
       REGION "COPY TO LOCAL"
           #selStnCount := #settings.current.stations.selCount;
       END_REGION

       REGION "ON CHANGE IN BUTTON OR STATION SELECTON"
           IF #settings.current.kp8.btnSelState <> #oldSelState OR #selStnCount <> #oldSelStnCount THEN

               REGION "COPY TO LOCAL"
                   #stnCount := #constants.stationCount - 1;
               END_REGION

               REGION "FOR SELECTED STATIONS"
                   FOR #i := 0 TO #stnCount DO
                       #stnSelected := #stations.current[#i].settings.selected;
                       IF #stnSelected THEN

                           REGION "SAVE BUTTON SELECTION STATE"
                               #stations.current[#i].settings.btnSelection := #settings.current.kp8.btnSelState;
                           END_REGION

                       END_IF;
                   END_FOR;
               END_REGION

           END_IF;
       END_REGION

       REGION "SELECTED STATION COUNT CHANGE DETECTION"
           #oldSelStnCount := #selStnCount; 
       END_REGION

   END_REGION

   REGION "COUNT SELECTED BUTTONS"

       REGION "COPY TO LOCAL"
           #btnCount := #constants.buttonCount - 1;
       END_REGION 

       REGION "ON CHANGE IN BUTTON SELECTION STATES"
           IF #settings.current.kp8.btnSelState <> #oldSelState THEN

               REGION "INITIALIZE LOCAL"
                   #count := 0;
               END_REGION

               REGION "FOR EACH SELECTED BUTTON"
                   FOR #i := 0 TO #btnCount DO
                       IF #settings.current.kp8.btnSelState[#i] THEN

                           REGION "INCREMENT COUNT"
                               #count := #count + 1;
                           END_REGION

                       END_IF;
                   END_FOR;
               END_REGION

               REGION "SAVE COUNT"
                   #settings.current.kp8.selCount := #count;
               END_REGION

           END_IF;
       END_REGION

   END_REGION 

   REGION "UI INTERACTION ANIMATIONS"

       REGION "SELECT ALL BUTTONS"
           #btnPress := #settings.current.kp8.selectButtons.actuate;
           #animate := "Animate Bool"(colorTrue := #constants.colorLib.BgLGr,
                                      colorFalse := #constants.colorLib.BgGray,
                                      evalSignal := #btnPress);
           #settings.current.kp8.selectButtons.animate := #animate;
       END_REGION

       REGION "STOP RESET SELECTED STATION"
           #btnPress := #settings.current.kp8.buttons[0].actuate;
           #animate := "Animate Bool"(colorTrue := #constants.colorLib.FgGray,
                                      colorFalse := #constants.colorLib.BgGray,
                                      evalSignal := #btnPress);
           #settings.current.kp8.buttons[0].animate := #animate;
       END_REGION

       REGION "STOP RUNTIME"
           #btnPress := #settings.current.kp8.buttons[4].actuate;
           #animate := "Animate Bool"(colorTrue := #constants.colorLib.FgGray,
                                      colorFalse := #constants.colorLib.BgGray,
                                      evalSignal := #btnPress);
           #settings.current.kp8.buttons[4].animate := #animate;
       END_REGION

       REGION "BUTTON SELECTIONS"

           REGION "COPY TO LOCAL"
               #btnCount := #constants.buttonCount - 1;
           END_REGION

           REGION "FOR EACH BUTTON"     
               FOR #i := 0 TO #btnCount DO

                   REGION "EXCLUDE STOP RUNTIME AND RESET SELECTED BUTTONS"
                       IF #i <> 0 AND #i <> 4 THEN

                           REGION "ANIMATE"

                               REGION "COPY TO LOCAL"
                                   #btnPress := #settings.current.kp8.buttons[#i].actuate;
                               END_REGION

                               REGION "ENABLE/DISABLE"
                                   #animate := "Animate Bool"(colorTrue := #constants.colorLib.BgGray,
                                                              colorFalse := #constants.colorLib.disabled,
                                                              evalSignal := #enableState);
                               END_REGION

                               REGION "ENABLED SUB ANIMATIONS"
                                   IF #enableState THEN

                                       REGION "BUTTON SELECTED"
                                           #animate := "Animate Bool"(colorTrue := #constants.colorLib.BgLTe,
                                                                      colorFalse := #animate,
                                                                      evalSignal := #settings.current.kp8.btnSelState[#i]);
                                       END_REGION

                                       REGION "BUTTON UP/DOWN"
                                           #animate := "Animate Bool"(colorTrue := #constants.colorLib.BgDTe,
                                                                      colorFalse := #animate,
                                                                      evalSignal := #btnPress);
                                       END_REGION
                                   END_IF;
                               END_REGION

                               REGION "SAVE ANIMATION"
                                   #settings.current.kp8.buttons[#i].animate := #animate;
                               END_REGION

                           END_REGION

                       END_IF;
                   END_REGION

               END_FOR;
           END_REGION

       END_REGION

   END_REGION

   REGION "DRAW KP8 BUTTON LABELS"
       IF #reset THEN
           #settings.current.kp8.buttons[1].label := wstring#'6';
           #settings.current.kp8.buttons[2].label := wstring#'4';
           #settings.current.kp8.buttons[3].label := wstring#'2';
           #settings.current.kp8.buttons[5].label := wstring#'5';
           #settings.current.kp8.buttons[6].label := wstring#'3';
           #settings.current.kp8.buttons[7].label := wstring#'1';
       END_IF;
   END_REGION

   REGION "CHANGE DETECTION"
       #oldSelState := #settings.current.kp8.btnSelState;
   END_REGION
END_FUNCTION_BLOCK

FUNCTION_BLOCK "Station Details"   // FB22, SCL
{ S7_Optimized_Access := 'TRUE' }
VERSION : 0.1
   VAR_INPUT
      constants : "Constants";
   END_VAR
   VAR_IN_OUT
      settings : "Settings Screen";
      stations : "Stations";
   END_VAR
   VAR
      old : Struct
         asgnPN : Bool;
         asgnAlloted : Bool;
         asgnCritical : Bool;
         nextPress : Bool;
         prevPress : Bool;
         selBtnCount : Int;
         selBtnNumber : Int;
         selStnCount : Int;
         selStnNumber : Int;
      END_STRUCT;
      selStnNumber : Int;
      selBtnNumber : Int;
      newViewReq : Bool;
      instPNEntEnable : "Enable Assignment Pair";
      instAlltEntEnable : "Enable Assignment Pair";
      instCrtEntEnable : "Enable Assignment Pair";
   END_VAR
   VAR_TEMP
      animate : USInt;
      btnCount : Int;
      btnPress : Bool;
      btnSelected : Bool;
      disable : Bool;
      dropZone : WString;
      enable : Bool;
      i : Int;
      j : Int;
      line : WString;
      partNumber : WString;
      pBtn : Int;
      selBtnCount : Int;
      selStnCount : Int;
      stnCount : Int;
      stnName : WString;
      stnSelected : Bool;
      timerWS : WString;
      timerReal : Real;
      labelEntered : Bool;
      lineLabel : WString;
      dzEntered : Bool;
      dzLabel : WString;
   END_VAR
   VAR CONSTANT
      blankString : WString;
   END_VAR
BEGIN
   REGION "POPULATE STATION NAME AND NUMBER"

       REGION "COPY TO LOCAL"
           #selStnCount := #settings.current.stations.selCount;
           #stnCount := #constants.stationCount - 1;
       END_REGION

       REGION "ON CHANGE IN STATION COUNT"
           IF #selStnCount <> #old.selStnCount AND #selStnCount <> 0 THEN

               REGION "FOR EACH STATION"
                   FOR #i := 0 TO #stnCount DO

                       REGION "COPY TO LOCAL"
                           #stnSelected := #stations.current[#i].settings.selected;
                       END_REGION

                       REGION "ON SELECTED STATION"
                           IF #stnSelected THEN

                               #selStnNumber := #i ;
                               EXIT;

                           END_IF;
                       END_REGION

                   END_FOR;
               END_REGION

           END_IF;
       END_REGION

   END_REGION

   REGION "PREVIOUS STATION"

       REGION "COPY TO LOCAL"
           #selStnCount := #settings.current.stations.selCount;
       END_REGION

       REGION "WHILE A STATION HAS BEEN SELECTED"
           IF #selStnCount <> 0 THEN

               REGION "COPY TO LOCAL"
                   #btnPress := #settings.current.viewingStation.previous.actuate;
                   #stnCount := #constants.stationCount - 1;
               END_REGION

               REGION "ON BUTTON PRESS RISING EDGE"
                   IF #btnPress AND NOT #old.prevPress THEN

                       REGION "INITIALIZE INDEX VARIABLE"
                           #i := #selStnNumber - 1;
                       END_REGION

                       REGION "LOW LIMIT ROLL OVER"
                           IF #i < 0 THEN
                               #i := #stnCount;
                           END_IF;
                       END_REGION

                       REGION "COPY TO LOCAL"
                           #stnSelected := #stations.current[#i].settings.selected;
                       END_REGION

                       REGION "FIND NEXT SELECTED STATION"
                           WHILE NOT #stnSelected DO

                               REGION "DECREMENT INDEX"
                                   #i -= 1;
                               END_REGION

                               REGION "EXIT LOOP NO STATION SELECTED"
                                   IF #i < 0 THEN
                                       #i := #stnCount;
                                   END_IF;
                               END_REGION

                               REGION "SAVE WHILE CONDITION"
                                   #stnSelected := #stations.current[#i].settings.selected;
                               END_REGION

                           END_WHILE;
                       END_REGION

                       REGION "SAVE NEW SELECTED STATION NUMBER"
                           #selStnNumber := #i;
                       END_REGION

                   END_IF;
               END_REGION

               REGION "CHANGE DETECTION"
                   #old.prevPress := #btnPress;
               END_REGION

           END_IF;
       END_REGION

   END_REGION

   REGION "NEXT STATION"

       REGION "COPY TO LOCAL"
           #selStnCount := #settings.current.stations.selCount;
       END_REGION

       REGION "WHILE A STATION HAS BEEN SELECTED"
           IF #selStnCount <> 0 THEN

               REGION "COPY TO LOCAL"
                   #btnPress := #settings.current.viewingStation.next.actuate;
                   #stnCount := #constants.stationCount - 1;
               END_REGION

               REGION "ON BUTTON PRESS RISING EDGE"
                   IF #btnPress AND NOT #old.nextPress OR #selStnCount <> #old.selStnCount THEN

                       REGION "INITIALIZE INDEX VARIABLE"
                           #i := #selStnNumber + 1;
                       END_REGION

                       REGION "LOW LIMIT ROLL OVER"
                           IF #i > #stnCount THEN
                               #i := 0;
                           END_IF;
                       END_REGION

                       REGION "COPY TO LOCAL"
                           #stnSelected := #stations.current[#i].settings.selected;
                       END_REGION

                       REGION "FIND NEXT SELECTED STATION"
                           WHILE NOT #stnSelected DO

                               REGION "DECREMENT INDEX"
                                   #i += 1;
                               END_REGION

                               REGION "EXIT LOOP NO STATION SELECTED"
                                   IF #i > #stnCount THEN
                                       #i := 0;
                                   END_IF;
                               END_REGION

                               REGION "SAVE WHILE CONDITION"
                                   #stnSelected := #stations.current[#i].settings.selected;
                               END_REGION

                           END_WHILE;
                       END_REGION

                       REGION "SAVE NEW SELECTED STATION NUMBER"
                           #selStnNumber := #i;
                       END_REGION

                   END_IF;
               END_REGION

               REGION "CHANGE DETECTION"
                   #old.nextPress := #btnPress;
               END_REGION

           END_IF;
       END_REGION


   END_REGION

   REGION "UPDATE STATION NAME"

       REGION "ON CHANGE IN SELECTED STAION NUMBER"
           IF #selStnNumber <> #old.selStnNumber THEN

               REGION "WRITE STATION NAME"
                   #line := #stations.current[#selStnNumber].line;
                   #dropZone := "Strip Sign"(USINT_TO_WSTRING(#stations.current[#selStnNumber].dropZone));
                   #stnName := CONCAT_WSTRING(IN1 := #line,
                                              IN2 := wstring#' ',
                                              IN3 := #dropZone);
                   #settings.current.viewingStation.name := #stnName;
               END_REGION

           END_IF;
       END_REGION



   END_REGION

   REGION "UPDATE LINE AND DROP ZONE DISPLAY"

       REGION "COPY TO LOCAL"
           #selStnCount := #settings.current.stations.selCount;
       END_REGION

       REGION "ON CHANGE IN SELECTED STAION NUMBER"
           IF #selStnCount <> #old.selStnCount AND #selStnCount = 1 THEN

               REGION "COPY TO LOCAL"
                   #line := #stations.current[#selStnNumber].line;
                   #dropZone := "Strip Sign"(USINT_TO_WSTRING(#stations.current[#selStnNumber].dropZone));
               END_REGION

               REGION "WRITE LINE AND DROP ZONE"
                   #settings.current.viewingStation.lineData.value := #line;
                   #settings.current.viewingStation.dzData.value := #dropZone;
               END_REGION

           END_IF;
       END_REGION



   END_REGION

   REGION "DISPLAY PN AND TIMER VALUES FOR BUTTON"

       REGION "COPY TO LOCAL"
           #selStnCount := #settings.current.stations.selCount;
           #selBtnCount := #settings.current.kp8.selCount;
           #selBtnNumber := #settings.current.kp8.selBtnNumber;
       END_REGION

       REGION "IF A STATION AND BUTTON HAVE BEEN SELECTED"
           IF #selStnCount <> 0 AND #selBtnCount <> 0 THEN

               REGION "ON NEW BUTTON SELECTION"
                   IF #selBtnCount <> #old.selBtnCount OR #selStnCount <> #old.selStnCount THEN

                       REGION "PART NUMBER"
                           #partNumber := #stations.current[#selStnNumber].partNumbers[#selBtnNumber];
                           #settings.current.partNumber.ioField.value := #partNumber;
                       END_REGION

                       REGION "ALLOTTED TIMER"
                           #timerWS := "Real to WString Timer"(#stations.current[#selStnNumber].presetTime.allotted[#selBtnNumber]);
                           #settings.current.alotted.ioField.value := #timerWS;
                       END_REGION

                       REGION "CRITITCAL TIMER"
                           #timerWS := "Real to WString Timer"(#stations.current[#selStnNumber].presetTime.critical[#selBtnNumber]);
                           #settings.current.critical.ioField.value := #timerWS;
                       END_REGION

                   END_IF;
               END_REGION

           END_IF;
       END_REGION

       REGION "ON NO SELECTION"
           IF #selStnCount = 0 OR #selBtnCount = 0 THEN

               REGION "PART NUMBER"
                   #settings.current.partNumber.ioField.value := #blankString;
               END_REGION

               REGION "ALLOTTED TIMER"
                   #settings.current.alotted.ioField.value := #blankString;
               END_REGION

               REGION "CRITITCAL TIMER"
                   #settings.current.critical.ioField.value := #blankString;
               END_REGION

           END_IF;
       END_REGION

   END_REGION

   REGION "ASSIGN VALUES TO STATION"

       REGION "PART NUMBER"

           REGION "COPY TO LOCAL"
               #btnPress := #settings.current.partNumber.assign.actuate;
               #stnCount := #constants.stationCount - 1;
               #btnCount := #constants.buttonCount - 1;
           END_REGION

           REGION "ON RISING EDGE"
               IF #btnPress AND NOT #old.asgnPN THEN

                   REGION "COPY TO LOCAL"
                       #partNumber := #settings.current.partNumber.ioField.value;
                   END_REGION

                   REGION "FOR EACH STATION"
                       FOR #i := 0 TO #stnCount DO

                           REGION "COPY TO LOCAL"
                               #stnSelected := #stations.current[#i].settings.selected;
                           END_REGION

                           REGION "ON SELECTED STATION"
                               IF #stnSelected THEN

                                   REGION "FOR EACH BUTTON"
                                       FOR #j := 0 TO #btnCount DO

                                           REGION "COPY TO LOCAL"
                                               #btnSelected := #stations.current[#i].settings.btnSelection[#j];
                                           END_REGION

                                           REGION "FOR EACH SELECTED BUTTON"
                                               IF #btnSelected THEN

                                                   REGION "ASSIGN PART NUMBER"
                                                       #stations.current[#i].partNumbers[#j] := #partNumber;
                                                   END_REGION

                                               END_IF;
                                           END_REGION

                                       END_FOR;
                                   END_REGION

                               END_IF;
                           END_REGION

                       END_FOR;
                   END_REGION

               END_IF;
           END_REGION


           REGION "CHANGE DETECTION"
               #old.asgnPN := #btnPress;
           END_REGION

       END_REGION

       REGION "ALLOTTED TIME"

           REGION "COPY TO LOCAL"
               #btnPress := #settings.current.alotted.assign.actuate;
               #stnCount := #constants.stationCount - 1;
               #btnCount := #constants.buttonCount - 1;
           END_REGION

           REGION "ON RISING EDGE"
               IF #btnPress AND NOT #old.asgnPN THEN

                   REGION "COPY TO LOCAL"
                       #timerReal := "WString Timer to Real"(#settings.current.alotted.ioField.value);
                   END_REGION

                   REGION "FOR EACH STATION"
                       FOR #i := 0 TO #stnCount DO

                           REGION "COPY TO LOCAL"
                               #stnSelected := #stations.current[#i].settings.selected;
                           END_REGION

                           REGION "ON SELECTED STATION"
                               IF #stnSelected THEN

                                   REGION "FOR EACH BUTTON"
                                       FOR #j := 0 TO #btnCount DO

                                           REGION "COPY TO LOCAL"
                                               #btnSelected := #stations.current[#i].settings.btnSelection[#j];
                                           END_REGION

                                           REGION "ON SELECTED BUTTON"
                                               IF #btnSelected THEN

                                                   REGION "ASSIGN TIMER VALUE"
                                                       #stations.current[#i].presetTime.allotted[#j] := #timerReal;
                                                   END_REGION

                                               END_IF;
                                           END_REGION

                                       END_FOR;
                                   END_REGION

                               END_IF;
                           END_REGION

                       END_FOR;
                   END_REGION

               END_IF;
           END_REGION


           REGION "CHANGE DETECTION"
               #old.asgnAlloted := #btnPress;
           END_REGION

       END_REGION

       REGION "CRITICAL TIME"

           REGION "COPY TO LOCAL"
               #btnPress := #settings.current.critical.assign.actuate;
               #stnCount := #constants.stationCount - 1;
               #btnCount := #constants.buttonCount - 1;
           END_REGION

           REGION "ON RISING EDGE"
               IF #btnPress AND NOT #old.asgnPN THEN

                   REGION "COPY TO LOCAL"                    
                       #timerReal := "WString Timer to Real"(#settings.current.critical.ioField.value);
                   END_REGION

                   REGION "FOR EACH STATION"
                       FOR #i := 0 TO #stnCount DO

                           REGION "COPY TO LOCAL"
                               #stnSelected := #stations.current[#i].settings.selected;
                           END_REGION

                           REGION "ON SELECTED STATION"
                               IF #stnSelected THEN

                                   REGION "FOR EACH BUTTON"
                                       FOR #j := 0 TO #btnCount DO

                                           REGION "COPY TO LOCAL"
                                               #btnSelected := #stations.current[#i].settings.btnSelection[#j];
                                           END_REGION

                                           REGION "ON SELECTED BUTTON"
                                               IF #btnSelected THEN

                                                   REGION "ASSIGN TIMER VALUE"
                                                       #stations.current[#i].presetTime.critical[#j] := #timerReal;
                                                   END_REGION

                                               END_IF;
                                           END_REGION

                                       END_FOR;
                                   END_REGION

                               END_IF;
                           END_REGION

                       END_FOR;
                   END_REGION

               END_IF;
           END_REGION


           REGION "CHANGE DETECTION"
               #old.asgnCritical := #btnPress;
           END_REGION


       END_REGION

       REGION "LINE LABEL"

           REGION "COPY TO LOCAL"
               #labelEntered := #settings.current.viewingStation.lineData.inputFinished;
               #stnCount := #constants.stationCount - 1;
           END_REGION

           REGION "ON RISING EDGE"
               IF #labelEntered THEN

                   REGION "TURN OFF THE LIGHTS"
                       #settings.current.viewingStation.lineData.inputFinished := FALSE;
                   END_REGION

                   REGION "COPY TO LOCAL"                    
                       #lineLabel := #settings.current.viewingStation.lineData.value;
                   END_REGION

                   REGION "FOR EACH STATION"
                       FOR #i := 0 TO #stnCount DO

                           REGION "COPY TO LOCAL"
                               #stnSelected := #stations.current[#i].settings.selected;
                           END_REGION

                           REGION "ON SELECTED STATION"
                               IF #stnSelected THEN

                                   REGION "ASSIGN TIMER VALUE"
                                       #stations.current[#i].line := #lineLabel;
                                   END_REGION

                               END_IF;
                           END_REGION

                       END_FOR;
                   END_REGION

               END_IF;
           END_REGION

       END_REGION

       REGION "DROP ZONE LABEL"

           REGION "COPY TO LOCAL"
               #dzEntered := #settings.current.viewingStation.dzData.inputFinished;
               #stnCount := #constants.stationCount - 1;
           END_REGION

           REGION "ON RISING EDGE"
               IF #dzEntered THEN

                   REGION "TURN OFF THE LIGHTS"
                       #settings.current.viewingStation.dzData.inputFinished := FALSE;
                   END_REGION

                   REGION "COPY TO LOCAL"                    
                       #dzLabel := #settings.current.viewingStation.dzData.value;
                   END_REGION

                   REGION "FOR EACH STATION"
                       FOR #i := 0 TO #stnCount DO

                           REGION "COPY TO LOCAL"
                               #stnSelected := #stations.current[#i].settings.selected;
                           END_REGION

                           REGION "ON SELECTED STATION"
                               IF #stnSelected THEN

                                   REGION "ASSIGN DROP ZONE VALUE"
                                       #stations.current[#i].dropZone := WSTRING_TO_USINT(#dzLabel);
                                   END_REGION

                               END_IF;
                           END_REGION

                       END_FOR;
                   END_REGION

               END_IF;
           END_REGION

       END_REGION

   END_REGION

   REGION "LOAD BUTTON DETAILS"

       REGION "COPY TO LOCAL"
           #selStnCount := #settings.current.stations.selCount;
           #btnCount := #constants.buttonCount - 3;
       END_REGION

       REGION "ON SELECTED STATIONS"
           IF #selStnCount >= 1 THEN

               REGION "FOR EACH BUTTON"
                   FOR #i := 0 TO #btnCount DO

                       REGION "CALCULATE BUTTON POINTER"
                           IF #i MOD 2 = 0 THEN
                               #pBtn := 7 - #i / 2;
                           END_IF;
                           IF #i MOD 2 <> 0 THEN
                               #pBtn := 3 - #i / 2;
                           END_IF;
                       END_REGION

                       REGION "BUTTON LABEL"
                           #settings.current.viewingStation.btns[#i].label.value := "Strip Sign"(INT_TO_WSTRING(#i + 1));
                       END_REGION

                       REGION "ALLOTTED TIME"
                           #timerWS := "Real to WString Timer"(#stations.current[#selStnNumber].presetTime.allotted[#pBtn]);
                           #settings.current.viewingStation.btns[#i].alloted.value := #timerWS;
                       END_REGION

                       REGION "CRITICAL TIME"
                           #timerWS := "Real to WString Timer"(#stations.current[#selStnNumber].presetTime.critical[#pBtn]);
                           #settings.current.viewingStation.btns[#i].critical.value := #timerWS;
                       END_REGION

                       REGION "PART NUMBER"
                           #partNumber := #stations.current[#selStnNumber].partNumbers[#pBtn];
                           #settings.current.viewingStation.btns[#i].partNumber.value := #partNumber;
                       END_REGION

                   END_FOR;
               END_REGION

           END_IF;
       END_REGION

   END_REGION

   REGION "ANIMATIONS"

       REGION "COPY TO LOCAL"
           #selStnCount := #settings.current.stations.selCount;
       END_REGION

       REGION "PN AND TIMERS"

           REGION "ENABLE/DISABLE FOR PN AND TIMERS"

               REGION "SET DISABLE"
                   IF #selStnCount = 0 OR #selBtnCount = 0 THEN
                       #disable := TRUE;
                       #enable := FALSE;
                   END_IF;
               END_REGION

               REGION "SET ENABLE"
                   IF #selStnCount <> 0 AND #selBtnCount <> 0 THEN
                       #disable := FALSE;
                       #enable := TRUE;
                   END_IF;
               END_REGION

           END_REGION

           REGION "PN ANIMATION FUNCTIONS"
               #animate := #settings.current.partNumber.assign.animate;
               #instPNEntEnable(constants := #constants,
                                disable := #disable,
                                enable := #enable,
                                value := #settings.current.partNumber.ioField.value,
                                assignAnimate := #animate,
                                ioFieldAnimate := #settings.current.partNumber.ioField.animate);
               #animate := "Animate Bool"(colorTrue := #constants.colorLib.BgLGr,
                                          colorFalse := #animate,
                                          evalSignal := #settings.current.partNumber.assign.actuate);
               #settings.current.partNumber.assign.animate := #animate;
           END_REGION

           REGION "ALLOTTED TIME ANIMATION FUNCTIONS"
               #animate := #settings.current.alotted.assign.animate;
               #instAlltEntEnable(constants := #constants,
                                  disable := #disable,
                                  enable := #enable,
                                  value := #settings.current.alotted.ioField.value,
                                  assignAnimate := #animate,
                                  ioFieldAnimate := #settings.current.alotted.ioField.animate);
               #animate := "Animate Bool"(colorTrue := #constants.colorLib.BgLGr,
                                          colorFalse := #animate,
                                          evalSignal := #settings.current.alotted.assign.actuate);
               #settings.current.alotted.assign.animate := #animate;
           END_REGION

           REGION "CRITICAL TIME ANIMATION FUNCTIONS"
               #animate := #settings.current.critical.assign.animate;
               #instCrtEntEnable(constants := #constants,
                                 disable := #disable,
                                 enable := #enable,
                                 value := #settings.current.critical.ioField.value,
                                 assignAnimate := #animate,
                                 ioFieldAnimate := #settings.current.critical.ioField.animate);
               #animate := "Animate Bool"(colorTrue := #constants.colorLib.BgLGr,
                                          colorFalse := #animate,
                                          evalSignal := #settings.current.critical.assign.actuate);
               #settings.current.critical.assign.animate := #animate;
           END_REGION

       END_REGION

       REGION "PREVIOUS STATION"
           #animate := "Animate Bool"(colorTrue := #constants.colorLib.BgLGr,
                                      colorFalse := #constants.colorLib.BgGray,
                                      evalSignal := #settings.current.viewingStation.previous.actuate);
           #settings.current.viewingStation.previous.animate := #animate;
       END_REGION

       REGION "NEXT STATION"
           #animate := "Animate Bool"(colorTrue := #constants.colorLib.BgLGr,
                                      colorFalse := #constants.colorLib.BgGray,
                                      evalSignal := #settings.current.viewingStation.next.actuate);
           #settings.current.viewingStation.next.animate := #animate;
       END_REGION

       REGION "ENABLE/DISABLE LINE DISPLAY"

           REGION "ENABLE"
               IF #selStnCount = 1 THEN
                   #settings.current.viewingStation.lineData.animate.bg := #constants.colorLib.BgGray;
                   #settings.current.viewingStation.lineData.animate.ioField := #constants.colorLib.BgWh;
               END_IF;
           END_REGION

           REGION "DISABLE"
               IF #selStnCount <> 1 THEN
                   #settings.current.viewingStation.lineData.animate.bg := #constants.colorLib.invisible;
                   #settings.current.viewingStation.lineData.animate.ioField := #constants.colorLib.invisible;
               END_IF;
           END_REGION

       END_REGION

       REGION "ENABLE/DISABLE DROPZONE"

           REGION "ENABLE"
               IF #selStnCount = 1 THEN
                   #settings.current.viewingStation.dzData.animate.bg := #constants.colorLib.BgGray;
                   #settings.current.viewingStation.dzData.animate.ioField := #constants.colorLib.BgWh;
               END_IF;
           END_REGION

           REGION "DISABLE"
               IF #selStnCount <> 1 THEN
                   #settings.current.viewingStation.dzData.animate.bg := #constants.colorLib.invisible;
                   #settings.current.viewingStation.dzData.animate.ioField := #constants.colorLib.invisible;
               END_IF;
           END_REGION

       END_REGION

       REGION "ENABLE/DISABLE BUTTON DETAILS"

           REGION "COPY TO LOCAL"
               #btnCount := #constants.buttonCount - 3;
           END_REGION

           REGION "ENABLE"
               IF #selStnCount >= 1 THEN

                   REGION "SHOW BUTTON DETAILS"
                       #animate := #constants.colorLib.BgGray;
                   END_REGION

               END_IF;
           END_REGION

           REGION "DISABLE"
               IF #selStnCount = 0 THEN

                   REGION "HIDE BUTTON DETAILS"
                       #animate := #constants.colorLib.invisible;
                   END_REGION

               END_IF;
           END_REGION

           REGION "APPLY ANIMATION"
               FOR #i := 0 TO #btnCount DO
                   #settings.current.viewingStation.btns[#i].label.animate := #animate;
                   #settings.current.viewingStation.btns[#i].alloted.animate := #animate;
                   #settings.current.viewingStation.btns[#i].critical.animate := #animate;
                   #settings.current.viewingStation.btns[#i].partNumber.animate := #animate;
               END_FOR;

           END_REGION 
       END_REGION

   END_REGION

   REGION "CHANGE DETECTION"
       #old.selStnNumber := #selStnNumber;
       #old.selBtnNumber := #selBtnNumber;
       #old.selBtnCount := #selBtnCount;
       #old.selStnCount := #selStnCount;
   END_REGION
END_FUNCTION_BLOCK

FUNCTION_BLOCK "Enable Assignment Pair"   // FB23, SCL
{ S7_Optimized_Access := 'TRUE' }
VERSION : 0.1
   VAR_INPUT
      constants : "Constants";
      disable : Bool;
      enable : Bool;
   END_VAR
   VAR_IN_OUT
      value : WString;
      assignAnimate : USInt;
      ioFieldAnimate : USInt;
   END_VAR
   VAR
      old : Struct
         disabled : Bool;
         enabled : Bool;
      END_STRUCT;
   END_VAR
BEGIN
   REGION "DISABLED"    
       IF #disable THEN
           #value := wstring#'';
           #assignAnimate := #constants.colorLib.disabled;
           #ioFieldAnimate := #constants.colorLib.disabled;
       END_IF;
   END_REGION

   REGION "ENABLED"
           IF #enable THEN
               #assignAnimate := #constants.colorLib.BgGray;
               #ioFieldAnimate := #constants.colorLib.BgWh;
           END_IF;
   END_REGION
END_FUNCTION_BLOCK

FUNCTION_BLOCK "KP8 Driver"   // FB101, SCL
{ S7_Optimized_Access := 'FALSE' }
VERSION : 0.1
   VAR_INPUT
      btnIn : Byte;   // byte that contains input data from kp8 buttons
      hardInit : Bool;   // initializes function. can be used for reset
      softInit : Bool;
      btn0Activate : Bool;   // true for on, false for off
      btn0Mode : Bool;   // true for maintained, false for momentary
      btn0Group : Int;
      btn0Flash : Bool;
      btn0ColorOn1 : String[10];   // enter: red OR green OR blue OR yellow OR white OR off
      btn0ColorOn2 : String[10];
      btn0ColorOff : String[10];   // enter: red OR green OR blue OR yellow OR white OR off
      btn1Activate : Bool;   // true for on, false for off
      btn1Mode : Bool;   // true for maintained, false for momentary
      btn1Group : Int;
      btn1Flash : Bool;
      btn1ColorOn1 : String[10];   // enter: red OR green OR blue OR yellow OR white OR off
      btn1ColorOn2 : String[10];
      btn1ColorOff : String[10];   // enter: red OR green OR blue OR yellow OR white OR off
      btn2Activate : Bool;   // true for on, false for off
      btn2Mode : Bool;   // true for maintained, false for momentary
      btn2Group : Int;
      btn2Flash : Bool;
      btn2ColorOn1 : String[10] := '';   // enter: red OR green OR blue OR yellow OR white OR off
      btn2ColorOn2 : String[10];
      btn2ColorOff : String[10];   // enter: red OR green OR blue OR yellow OR white OR off
      btn3Activate : Bool;   // true for on, false for off
      btn3Mode : Bool;   // true for maintained, false for momentary
      btn3Group : Int;
      btn3Flash : Bool;
      btn3ColorOn1 : String[10];   // enter: red OR green OR blue OR yellow OR white OR off
      btn3ColorOn2 : String[10];
      btn3ColorOff : String[10];   // enter: red OR green OR blue OR yellow OR white OR off
      btn4Activate : Bool;   // true for on, false for off
      btn4Mode : Bool;   // true for maintained, false for momentary
      btn4Group : Int;
      btn4Flash : Bool;
      btn4ColorOn1 : String[10];   // enter: red OR green OR blue OR yellow OR white OR off
      btn4ColorOn2 : String[10];
      btn4ColorOff : String[10];   // enter: red OR green OR blue OR yellow OR white OR off
      btn5Activate : Bool;   // true for on, false for off
      btn5Mode : Bool;   // true for maintained, false for momentary
      btn5Group : Int;
      btn5Flash : Bool;
      btn5ColorOn1 : String[10];   // enter: red OR green OR blue OR yellow OR white OR off
      btn5ColorOn2 : String[10];
      btn5ColorOff : String[10];   // enter: red OR green OR blue OR yellow OR white OR off
      btn6Activate : Bool;   // true for on, false for off
      btn6Mode : Bool;   // true for maintained, false for momentary
      btn6Group : Int;
      btn6Flash : Bool;
      btn6ColorOn1 : String[10];   // enter: red OR green OR blue OR yellow OR white OR off
      btn6ColorOn2 : String[10];
      btn6ColorOff : String[10];   // enter: red OR green OR blue OR yellow OR white OR off
      btn7Activate : Bool;   // true for on, false for off
      btn7Mode : Bool;   // true for maintained, false for momentary
      btn7Group : Int;
      btn7Flash : Bool;
      btn7ColorOn1 : String[10];   // enter: red OR green OR blue OR yellow OR white OR off
      btn7ColorOn2 : String[10];
      btn7ColorOff : String[10];   // enter: red OR green OR blue OR yellow OR white OR off
   END_VAR
   VAR_OUTPUT
      btnStatesOut : Array[0..7] of Bool;   // the output array represents the state of button presses
      btnColorsOut : DWord;
   END_VAR
   VAR
      mask : Byte;
      btnInInt : Byte;
      btnEval : Byte;
      i1 : Int;
      i2 : Int;
      btnInArrayNew : Array[0..7] of Bool;
      btnInArrayOld : Array[0..7] of Bool;
      btnStateArrayInt : Array[0..7] of Bool;
      btnActivateInt : Array[0..7] of Bool;
      btnModeInt : Array[0..7] of Bool;
      btnFlashInt : Array[0..7] of Bool;
      btnGroup : Array[0..7] of Int;
      btnClrMskOn1Int : Array[0..7] of DWord;
      btnClrMskOn2Int : Array[0..7] of DWord;
      btnClrMskOffInt : Array[0..7] of DWord;
      btnClrOn1Int : Array[0..7] of String[10];
      btnClrOn2Int : Array[0..7] of String[10];
      btnClrOffInt : Array[0..7] of String[10];
   END_VAR
   VAR CONSTANT
      btnMskRed : DWord := dw#16#0100_0000;
      btnMskGreen : DWord := dw#16#0001_0000;
      btnMskBlue : DWord := dw#16#000_0100;
      btnMskYellow : DWord := dw#16#0101_0000;
      btnMskWhite : DWord := dw#16#0101_0100;
      btnMskBlack : DWord := dw#16#FEFE_FEFF;
      initBtnColors : DWord := dw#16#0000_0000;
   END_VAR
BEGIN
   REGION "ALL INITS"
       IF #hardInit OR #softInit THEN

           REGION "CLEAR OUTPUT COLORS"
               #btnColorsOut := #initBtnColors;
           END_REGION

           REGION "TRANSFER PARAMETERS TO INTERNAL ARRAYS"

               REGION "BUTTON 0"
                   #btnActivateInt[0] := #btn0Activate;
                   #btnModeInt[0] := #btn0Mode;
                   #btnGroup[0] := #btn0Group;
                   #btnClrOn1Int[0] := #btn0ColorOn1;
                   #btnClrOn2Int[0] := #btn0ColorOn2;
                   #btnClrOffInt[0] := #btn0ColorOff;
               END_REGION

               REGION "BUTTON 1"
                   #btnActivateInt[1] := #btn1Activate;
                   #btnModeInt[1] := #btn1Mode;
                   #btnGroup[1] := #btn1Group;
                   #btnClrOn1Int[1] := #btn1ColorOn1;
                   #btnClrOn2Int[1] := #btn1ColorOn2;
                   #btnClrOffInt[1] := #btn1ColorOff;
               END_REGION

               REGION "BUTTON 2"
                   #btnActivateInt[2] := #btn2Activate;
                   #btnModeInt[2] := #btn2Mode;
                   #btnGroup[2] := #btn2Group;
                   #btnClrOn1Int[2] := #btn2ColorOn1;
                   #btnClrOn2Int[2] := #btn2ColorOn2;
                   #btnClrOffInt[2] := #btn2ColorOff;
               END_REGION

               REGION "BUTTON 3"
                   #btnActivateInt[3] := #btn3Activate;
                   #btnModeInt[3] := #btn3Mode;
                   #btnGroup[3] := #btn3Group;
                   #btnClrOn1Int[3] := #btn3ColorOn1;
                   #btnClrOn2Int[3] := #btn3ColorOn2;
                   #btnClrOffInt[3] := #btn3ColorOff;
               END_REGION

               REGION "BUTTON 4"
                   #btnActivateInt[4] := #btn4Activate;
                   #btnModeInt[4] := #btn4Mode;
                   #btnGroup[4] := #btn4Group;
                   #btnClrOn1Int[4] := #btn4ColorOn1;
                   #btnClrOn2Int[4] := #btn4ColorOn2;
                   #btnClrOffInt[4] := #btn4ColorOff;
               END_REGION

               REGION "BUTTON 5"
                   #btnActivateInt[5] := #btn5Activate;
                   #btnModeInt[5] := #btn5Mode;
                   #btnGroup[5] := #btn5Group;
                   #btnClrOn1Int[5] := #btn5ColorOn1;
                   #btnClrOn2Int[5] := #btn5ColorOn2;
                   #btnClrOffInt[5] := #btn5ColorOff;
               END_REGION

               REGION "BUTTON 6"
                   #btnActivateInt[6] := #btn6Activate;
                   #btnModeInt[6] := #btn6Mode;
                   #btnGroup[6] := #btn6Group;
                   #btnClrOn1Int[6] := #btn6ColorOn1;
                   #btnClrOn2Int[6] := #btn6ColorOn2;
                   #btnClrOffInt[6] := #btn6ColorOff;
               END_REGION

               REGION "BUTTON 7"
                   #btnActivateInt[7] := #btn7Activate;
                   #btnModeInt[7] := #btn7Mode;
                   #btnGroup[7] := #btn7Group;
                   #btnClrOn1Int[7] := #btn7ColorOn1;
                   #btnClrOn2Int[7] := #btn7ColorOn2;
                   #btnClrOffInt[7] := #btn7ColorOff;
               END_REGION

           END_REGION

           REGION "RECOLOR BUTTON MASKS"
               FOR #i1 := 0 TO 7 DO

                   REGION "ON COLOR 1"
                       IF (#btnClrOn1Int[#i1] = 'red') THEN
                           #btnClrMskOn1Int[#i1] := SHL(IN := #btnMskRed, N := #i1);
                       ELSIF (#btnClrOn1Int[#i1] = 'green') THEN
                           #btnClrMskOn1Int[#i1] := SHL(IN := #btnMskGreen, N := #i1);
                       ELSIF (#btnClrOn1Int[#i1] = 'blue') THEN
                           #btnClrMskOn1Int[#i1] := SHL(IN := #btnMskBlue, N := #i1);
                       ELSIF (#btnClrOn1Int[#i1] = 'yellow') THEN
                           #btnClrMskOn1Int[#i1] := SHL(IN := #btnMskYellow, N := #i1);
                       ELSIF (#btnClrOn1Int[#i1] = 'white') THEN
                           #btnClrMskOn1Int[#i1] := SHL(IN := #btnMskWhite, N := #i1);
                       ELSIF (#btnClrOn1Int[#i1] = 'off') THEN
                           #btnClrMskOn1Int[#i1] := 0;
                       END_IF;
                   END_REGION

                   REGION "ON COLOR 2"
                       IF (#btnClrOn2Int[#i1] = 'red') THEN
                           #btnClrMskOn2Int[#i1] := SHL(IN := #btnMskRed, N := #i1);
                       ELSIF (#btnClrOn2Int[#i1] = 'green') THEN
                           #btnClrMskOn2Int[#i1] := SHL(IN := #btnMskGreen, N := #i1);
                       ELSIF (#btnClrOn2Int[#i1] = 'blue') THEN
                           #btnClrMskOn2Int[#i1] := SHL(IN := #btnMskBlue, N := #i1);
                       ELSIF (#btnClrOn2Int[#i1] = 'yellow') THEN
                           #btnClrMskOn2Int[#i1] := SHL(IN := #btnMskYellow, N := #i1);
                       ELSIF (#btnClrOn2Int[#i1] = 'white') THEN
                           #btnClrMskOn2Int[#i1] := SHL(IN := #btnMskWhite, N := #i1);
                       ELSIF (#btnClrOn2Int[#i1] = 'off') THEN
                           #btnClrMskOn2Int[#i1] := 0;
                       END_IF;
                   END_REGION

                   REGION "OFF COLOR"
                       IF (#btnClrOffInt[#i1] = 'red') THEN
                           #btnClrMskOffInt[#i1] := SHL(IN := #btnMskRed, N := #i1);
                       ELSIF (#btnClrOffInt[#i1] = 'green') THEN
                           #btnClrMskOffInt[#i1] := SHL(IN := #btnMskGreen, N := #i1);
                       ELSIF (#btnClrOffInt[#i1] = 'blue') THEN
                           #btnClrMskOffInt[#i1] := SHL(IN := #btnMskBlue, N := #i1);
                       ELSIF (#btnClrOffInt[#i1] = 'yellow') THEN
                           #btnClrMskOffInt[#i1] := SHL(IN := #btnMskYellow, N := #i1);
                       ELSIF (#btnClrOffInt[#i1] = 'white') THEN
                           #btnClrMskOffInt[#i1] := SHL(IN := #btnMskWhite, N := #i1);
                       ELSIF (#btnClrOffInt[#i1] = 'off') THEN
                           #btnClrMskOffInt[#i1] := 0;
                       END_IF;
                   END_REGION

               END_FOR;
           END_REGION

       END_IF;
   END_REGION

   REGION "HART INIT"
       IF #hardInit THEN
           FOR #i1 := 0 TO 7 DO
               #btnStateArrayInt[#i1] := FALSE;
           END_FOR;
       END_IF;
   END_REGION


   REGION "TRANFER PARAMETERS TO ARRAYS"
       // raw pb data
       #btnInInt := #btnIn;
       // flashing modes
       #btnFlashInt[0] := #btn0Flash;
       #btnFlashInt[1] := #btn1Flash;
       #btnFlashInt[2] := #btn2Flash;
       #btnFlashInt[3] := #btn3Flash;
       #btnFlashInt[4] := #btn4Flash;
       #btnFlashInt[5] := #btn5Flash;
       #btnFlashInt[6] := #btn6Flash;
       #btnFlashInt[7] := #btn7Flash;
   END_REGION

   REGION "EVALUATE BUTTONS"
       FOR #i1 := 0 TO 7 DO

           REGION "TRANSFER BUTTON PRESSES TO ARRAY"
               #btnEval := SHR(IN := #btnInInt, N := #i1);
               #btnInArrayNew[#i1] := #btnEval.%X0;
               #btnEval := b#16#0;
           END_REGION

           REGION "SET BUTTON STATE"

               REGION "BUTTON ACTIVE"
                   IF #btnActivateInt[#i1] THEN

                       REGION "MAINTAINED"
                           IF #btnModeInt[#i1] THEN

                               REGION "RISING EDGE OF PRESS"
                                   IF #btnInArrayNew[#i1] AND NOT #btnInArrayOld[#i1] THEN

                                       REGION "CHECK FOR GROUP MEMBERSHIP"
                                           FOR #i2 := 0 TO 7 DO

                                               REGION "NOT IN NULL GROUP"
                                                   IF (#btnGroup[#i2] <> 0) THEN

                                                       REGION "SKIP SELF"
                                                           IF (#i2 <> #i1) THEN

                                                               REGION "GROUPS MATCH"
                                                                   IF #btnGroup[#i1] = #btnGroup[#i2] THEN
                                                                       REGION "DEACTIVATE OTHER GROUP MEMBERS"
                                                                           #btnStateArrayInt[#i2] := FALSE;
                                                                       END_REGION

                                                                   END_IF;
                                                               END_REGION

                                                           END_IF;
                                                       END_REGION

                                                   END_IF;
                                               END_REGION

                                           END_FOR;
                                       END_REGION

                                       REGION "TOGGLE STATE"
                                           #btnStateArrayInt[#i1] := NOT #btnStateArrayInt[#i1];
                                       END_REGION

                                   END_IF;
                               END_REGION

                           END_IF;
                       END_REGION

                       REGION "MOMENTARY"
                           IF NOT #btnModeInt[#i1] THEN
                               #btnStateArrayInt[#i1] := #btnInArrayNew[#i1];
                           END_IF;
                       END_REGION

                   END_IF;
               END_REGION

               REGION "BUTTON INACTIVE"
                   IF NOT #btnActivateInt[#i1] THEN
                       #btnStateArrayInt[#i1] := FALSE;
                   END_IF;
               END_REGION

           END_REGION

           REGION "ANIMATE BUTTONS"

               REGION "BUTTON ON FLASH BIT OFF"
                   IF #btnStateArrayInt[#i1] AND NOT #btnFlashInt[#i1] THEN
                       #btnColorsOut := #btnColorsOut AND ROL(IN := #btnMskBlack, N := #i1);
                       #btnColorsOut := #btnColorsOut OR #btnClrMskOn1Int[#i1];
                   END_IF;
               END_REGION

